(* Logix 5000 project; controller FV vendor 1 type 14 code 217 rev 31.11; software revision 31.00; part 13 of 63 *)
(* tags used below, declared in another part *)
   CWD : CHECKWORD_FLAGS;
   FR_B240 : INT[255];   // DEBOUNCE Debounce Flags
   FR_B246 : INT[255];   // V_REVERSE Flags for reversing contol action
   FR_B3 : INT[255];   // BINARY
   FR_FV29_AV01 : PlantItem;   // FV29_AV01
   FR_FV29_AV04 : PlantItem;   // FV29_AV04
   FR_FV29_AV05 : PlantItem;   // FV29_AV05
   FR_FV29_AV06 : PlantItem;   // FV29_AV06
   FR_FV29_AV07 : PlantItem;   // FV29_AV07
   FR_FV29_ROTO : PlantItem;   // FV29_ROTO
   FR_FV29_VA01 : PlantItem;   // FV29_VA01
   FR_FV30_AV01 : PlantItem;   // FV30_AV01
   FR_FV30_AV04 : PlantItem;   // FV30_AV04
   FR_FV30_AV05 : PlantItem;   // FV30_AV05
   FR_FV30_AV06 : PlantItem;   // FV30_AV06
   FR_FV30_AV07 : PlantItem;   // FV30_AV07
   FR_FV30_ROTO : PlantItem;   // FV30_ROTO
   FR_FV30_VA01 : PlantItem;   // FV30_VA01
   FR_N10 : INT[265];   // FV_AGING Comms to FV Aging PL C
   FR_N100 : INT[265];   // FV FILLING
   FR_N110 : INT[265];   // GREEN BEER Green Beer Main
   FR_N120 : INT[265];   // YEAST CROP Yeast Cropping Main
   FR_N13 : INT[265];   // MV_ROUTE Comms to MV Routing PLC
   FR_N130 : INT[265];   // FILTRATE Filtrate Return
   FR_N14 : INT[265];   // MVFV CIP Comms to MVFV CIP Un it PLC
   FR_N160 : INT[265];   // VESSEL Vessel Working Direc tory
   FR_N200 : INT[265];   // ANALOG_IN Analog Inputs
   FR_N255 : INT[265];   // CHECKWORDS
   FR_N29 : INT[265];   // FV29
   FR_N30 : INT[265];   // FV30
   FR_N7 : INT[265];   // INTEGER
   FR_N99 : INT[265];   // COMMENT Comment Lines
   FR_T144 : TIMER[255];   // CIP
   FR_T4 : TIMER[255];   // TIMER
   FR_T50 : TIMER[52];
   FR_T51 : TIMER[52];
   FR_T52 : TIMER[52];
   FR_T53 : TIMER[52];
   FR_VB1_AV08 : PlantItem;   // VB1_AV08
   FR_VB1_AV09 : PlantItem;   // VB1_AV09
   FR_VB2_AV04 : PlantItem;   // VB2_AV04
   FR_VB2_AV05 : PlantItem;   // VB2_AV05
   FR_VB3_AV04 : PlantItem;   // VB3_AV04
   FR_VB3_AV05 : PlantItem;   // VB3_AV05
   FR_VB4_AV04 : PlantItem;   // VB4_AV04
   FR_VB4_AV05 : PlantItem;   // VB4_AV05
   FR_VB4_AV10 : PlantItem;   // VB4_AV10
   FR_VB4_AV11 : PlantItem;   // VB4_AV11
   FR_VB4_AV16 : PlantItem;   // VB4_AV16
   FR_VB4_AV17 : PlantItem;   // VB4_AV17
(* FR_Common, continued *)

ROUTINE FR_FV29_29   (* ladder *)
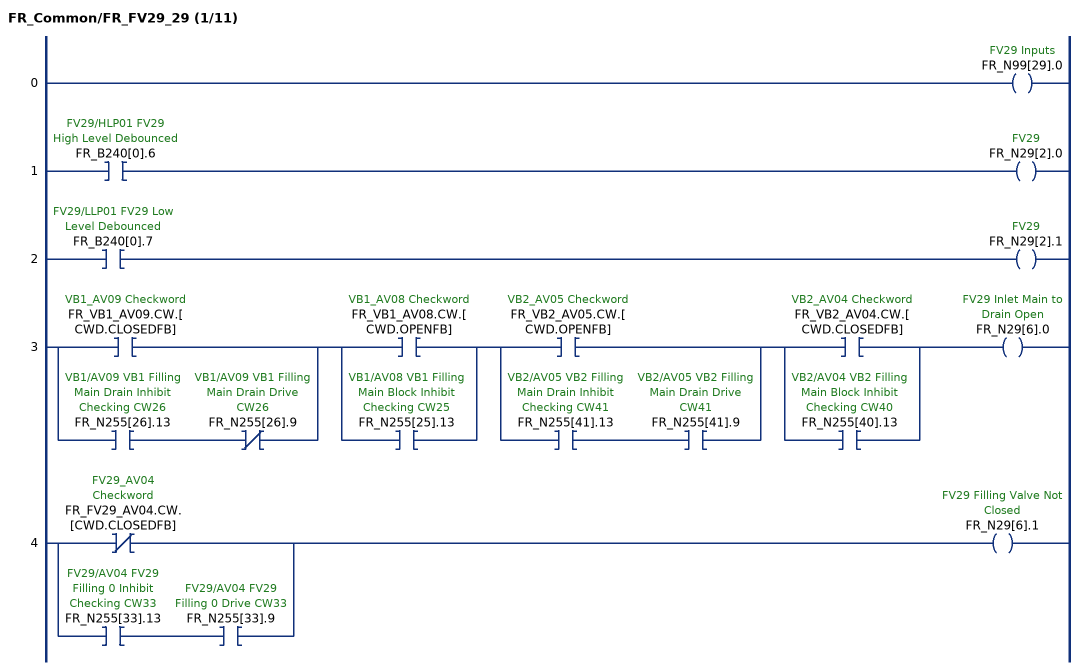
   0: OTE(FR_N99[29].0);
   1: XIC(FR_B240[0].6)OTE(FR_N29[2].0);
   2: XIC(FR_B240[0].7)OTE(FR_N29[2].1);
   3: [XIC(FR_VB1_AV09.CW.[CWD.CLOSEDFB]) ,XIC(FR_N255[26].13) XIO(FR_N255[26].9) ][XIC(FR_VB1_AV08.CW.[CWD.OPENFB]) ,XIC(FR_N255[25].13) ][XIC(FR_VB2_AV05.CW.[CWD.OPENFB]) ,XIC(FR_N255[41].13) XIC(FR_N255[41].9) ][XIC(FR_VB2_AV04.CW.[CWD.CLOSEDFB]) ,XIC(FR_N255[40].13) ]OTE(FR_N29[6].0);
   4: [XIO(FR_FV29_AV04.CW.[CWD.CLOSEDFB]) ,XIC(FR_N255[33].13) XIC(FR_N255[33].9) ]OTE(FR_N29[6].1);
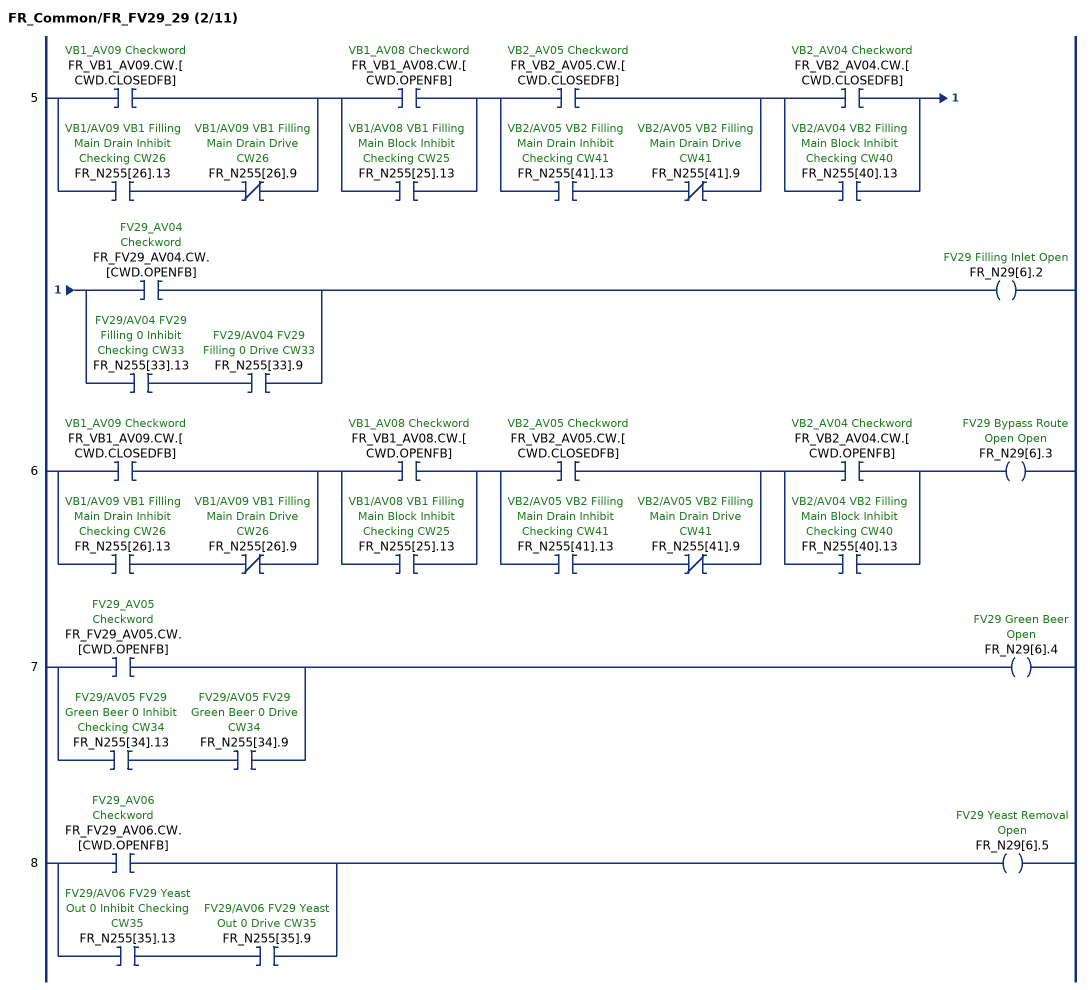
   5: [XIC(FR_VB1_AV09.CW.[CWD.CLOSEDFB]) ,XIC(FR_N255[26].13) XIO(FR_N255[26].9) ][XIC(FR_VB1_AV08.CW.[CWD.OPENFB]) ,XIC(FR_N255[25].13) ][XIC(FR_VB2_AV05.CW.[CWD.CLOSEDFB]) ,XIC(FR_N255[41].13) XIO(FR_N255[41].9) ][XIC(FR_VB2_AV04.CW.[CWD.CLOSEDFB]) ,XIC(FR_N255[40].13) ][XIC(FR_FV29_AV04.CW.[CWD.OPENFB]) ,XIC(FR_N255[33].13) XIC(FR_N255[33].9) ]OTE(FR_N29[6].2);
   6: [XIC(FR_VB1_AV09.CW.[CWD.CLOSEDFB]) ,XIC(FR_N255[26].13) XIO(FR_N255[26].9) ][XIC(FR_VB1_AV08.CW.[CWD.OPENFB]) ,XIC(FR_N255[25].13) ][XIC(FR_VB2_AV05.CW.[CWD.CLOSEDFB]) ,XIC(FR_N255[41].13) XIO(FR_N255[41].9) ][XIC(FR_VB2_AV04.CW.[CWD.OPENFB]) ,XIC(FR_N255[40].13) ]OTE(FR_N29[6].3);
   7: [XIC(FR_FV29_AV05.CW.[CWD.OPENFB]) ,XIC(FR_N255[34].13) XIC(FR_N255[34].9) ]OTE(FR_N29[6].4);
   8: [XIC(FR_FV29_AV06.CW.[CWD.OPENFB]) ,XIC(FR_N255[35].13) XIC(FR_N255[35].9) ]OTE(FR_N29[6].5);
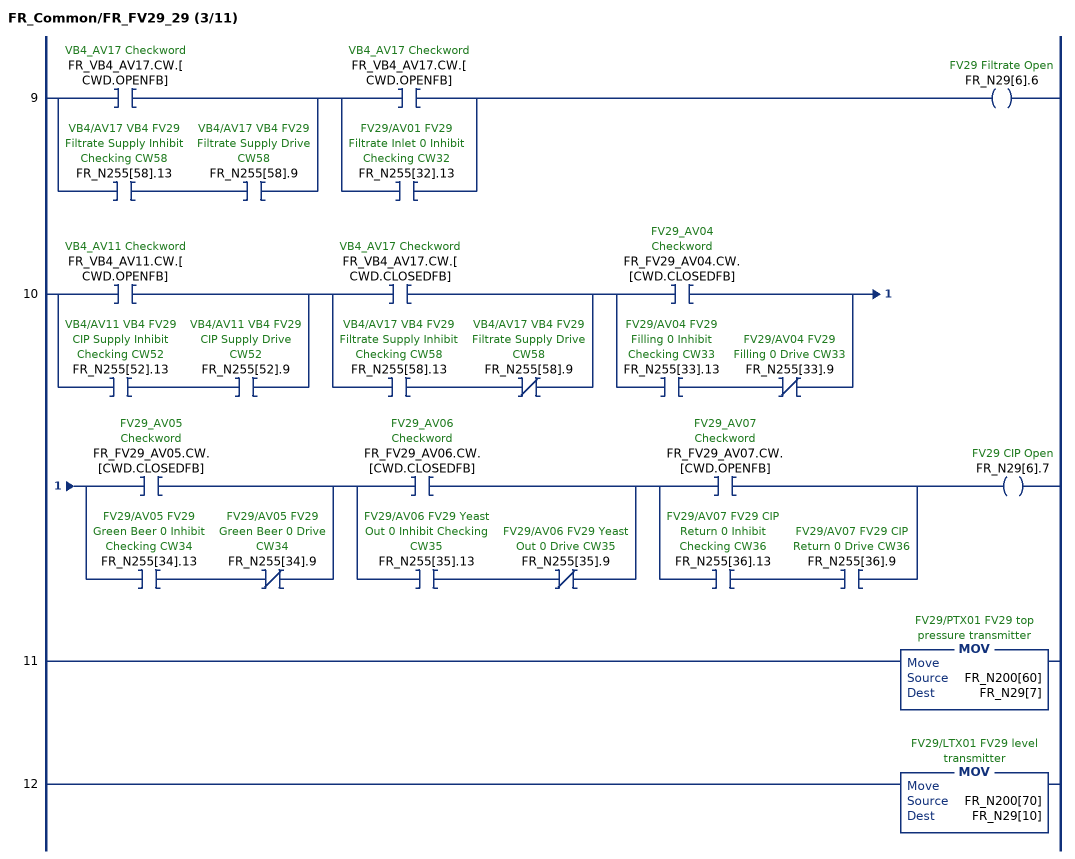
   9: [XIC(FR_VB4_AV17.CW.[CWD.OPENFB]) ,XIC(FR_N255[58].13) XIC(FR_N255[58].9) ][XIC(FR_VB4_AV17.CW.[CWD.OPENFB]) ,XIC(FR_N255[32].13) ]OTE(FR_N29[6].6);
   10: [XIC(FR_VB4_AV11.CW.[CWD.OPENFB]) ,XIC(FR_N255[52].13) XIC(FR_N255[52].9) ][XIC(FR_VB4_AV17.CW.[CWD.CLOSEDFB]) ,XIC(FR_N255[58].13) XIO(FR_N255[58].9) ][XIC(FR_FV29_AV04.CW.[CWD.CLOSEDFB]) ,XIC(FR_N255[33].13) XIO(FR_N255[33].9) ][XIC(FR_FV29_AV05.CW.[CWD.CLOSEDFB]) ,XIC(FR_N255[34].13) XIO(FR_N255[34].9) ][XIC(FR_FV29_AV06.CW.[CWD.CLOSEDFB]) ,XIC(FR_N255[35].13) XIO(FR_N255[35].9) ][XIC(FR_FV29_AV07.CW.[CWD.OPENFB]) ,XIC(FR_N255[36].13) XIC(FR_N255[36].9) ]OTE(FR_N29[6].7);
   11: MOV(FR_N200[60],FR_N29[7]);
   12: MOV(FR_N200[70],FR_N29[10]);
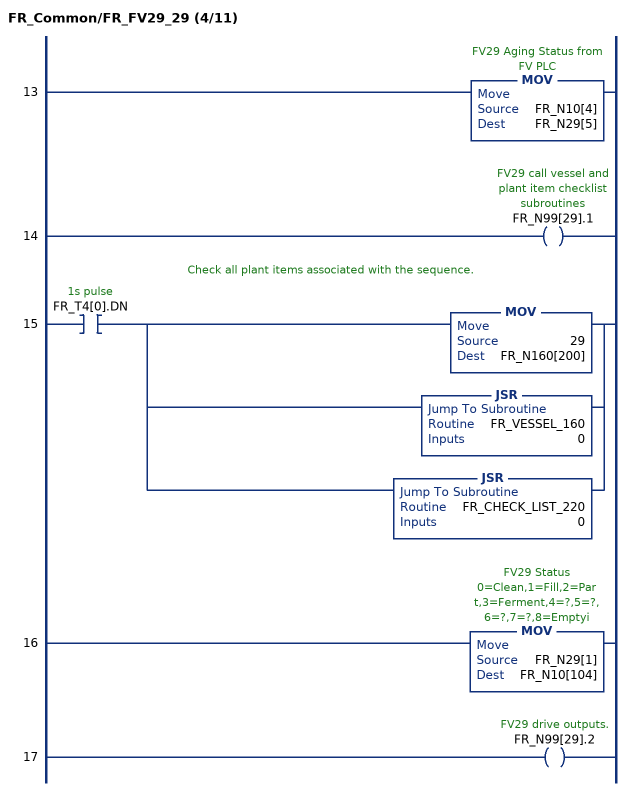
   13: MOV(FR_N10[4],FR_N29[5]);
   14: OTE(FR_N99[29].1);
   // Check all plant items associated with the sequence.
   15: XIC(FR_T4[0].DN)[MOV(29,FR_N160[200]) ,JSR(FR_VESSEL_160,0) ,JSR(FR_CHECK_LIST_220,0) ];
   16: MOV(FR_N29[1],FR_N10[104]);
   17: OTE(FR_N99[29].2);
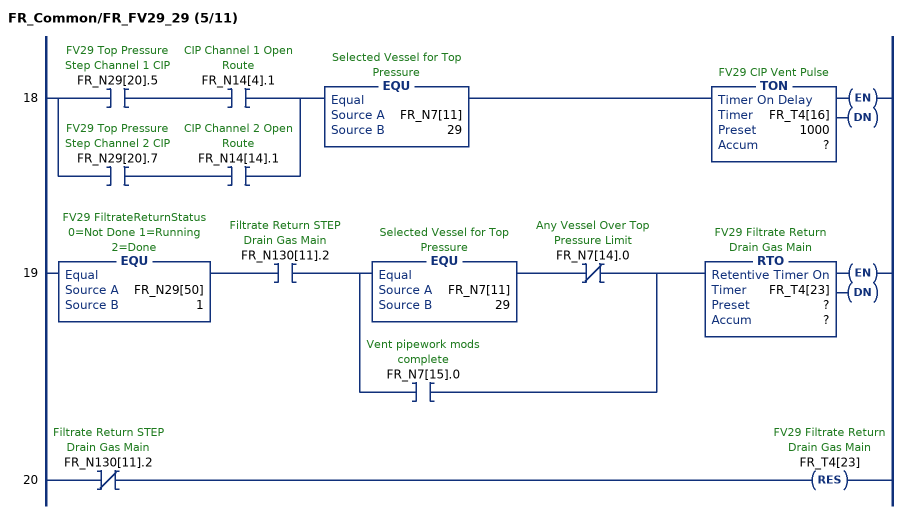
   18: [XIC(FR_N29[20].5) XIC(FR_N14[4].1) ,XIC(FR_N29[20].7) XIC(FR_N14[14].1) ]EQU(FR_N7[11],29)TON(FR_T4[16],?,?);
   19: EQU(FR_N29[50],1)XIC(FR_N130[11].2)[EQU(FR_N7[11],29) XIO(FR_N7[14].0) ,XIC(FR_N7[15].0) ]RTO(FR_T4[23],?,?);
   20: XIO(FR_N130[11].2)RES(FR_T4[23]);
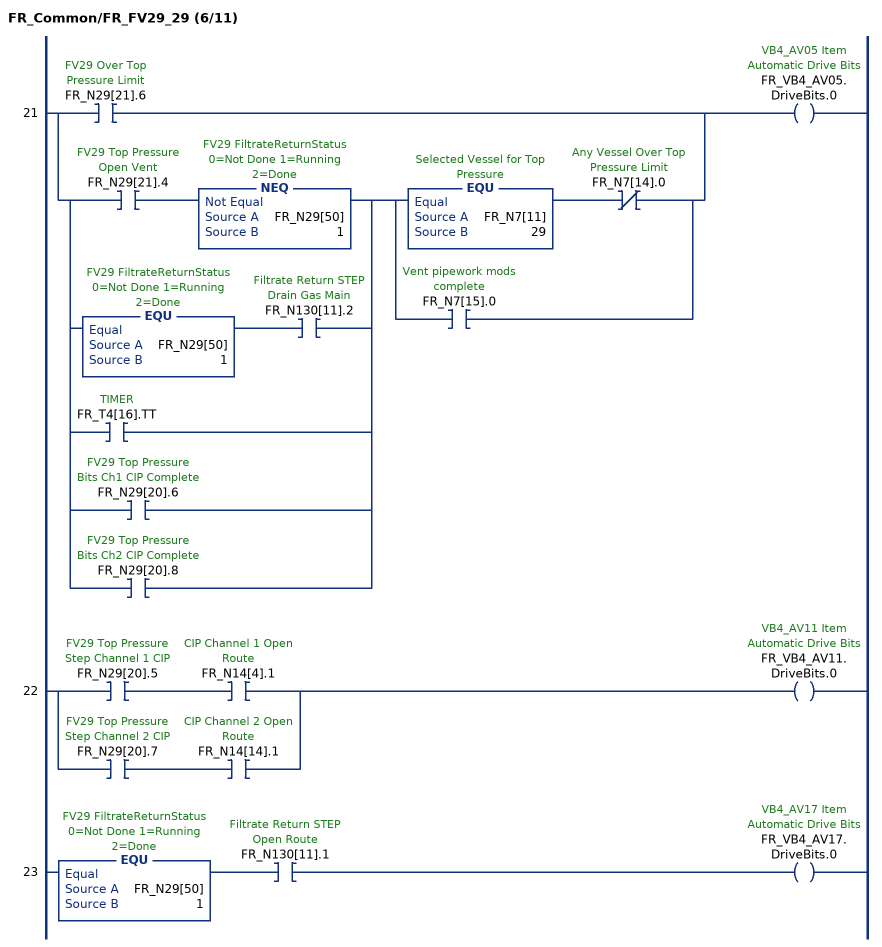
   21: [XIC(FR_N29[21].6) ,[XIC(FR_N29[21].4) NEQ(FR_N29[50],1) ,EQU(FR_N29[50],1) XIC(FR_N130[11].2) ,XIC(FR_T4[16].TT) ,[XIC(FR_N29[20].6) ,XIC(FR_N29[20].8) ] ] [EQU(FR_N7[11],29) XIO(FR_N7[14].0) ,XIC(FR_N7[15].0) ] ]OTE(FR_VB4_AV05.DriveBits.0);
   22: [XIC(FR_N29[20].5) XIC(FR_N14[4].1) ,XIC(FR_N29[20].7) XIC(FR_N14[14].1) ]OTE(FR_VB4_AV11.DriveBits.0);
   23: EQU(FR_N29[50],1)XIC(FR_N130[11].1)OTE(FR_VB4_AV17.DriveBits.0);
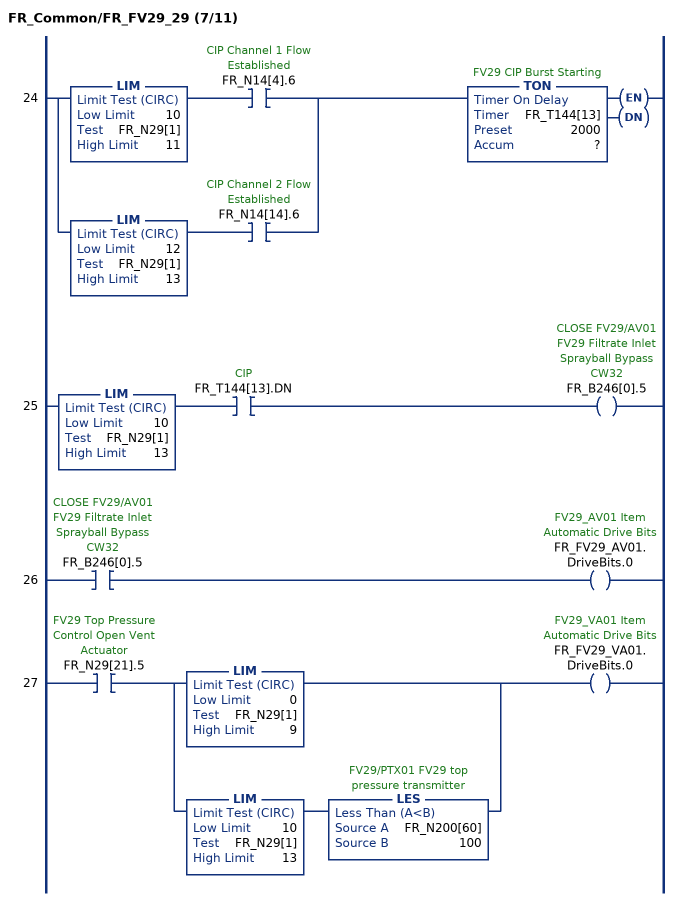
   24: [LIM(10,FR_N29[1],11) XIC(FR_N14[4].6) ,LIM(12,FR_N29[1],13) XIC(FR_N14[14].6) ]TON(FR_T144[13],?,?);
   25: LIM(10,FR_N29[1],13)XIC(FR_T144[13].DN)OTE(FR_B246[0].5);
   26: XIC(FR_B246[0].5)OTE(FR_FV29_AV01.DriveBits.0);
   27: XIC(FR_N29[21].5)[LIM(0,FR_N29[1],9) ,LIM(10,FR_N29[1],13) LES(FR_N200[60],100) ]OTE(FR_FV29_VA01.DriveBits.0);
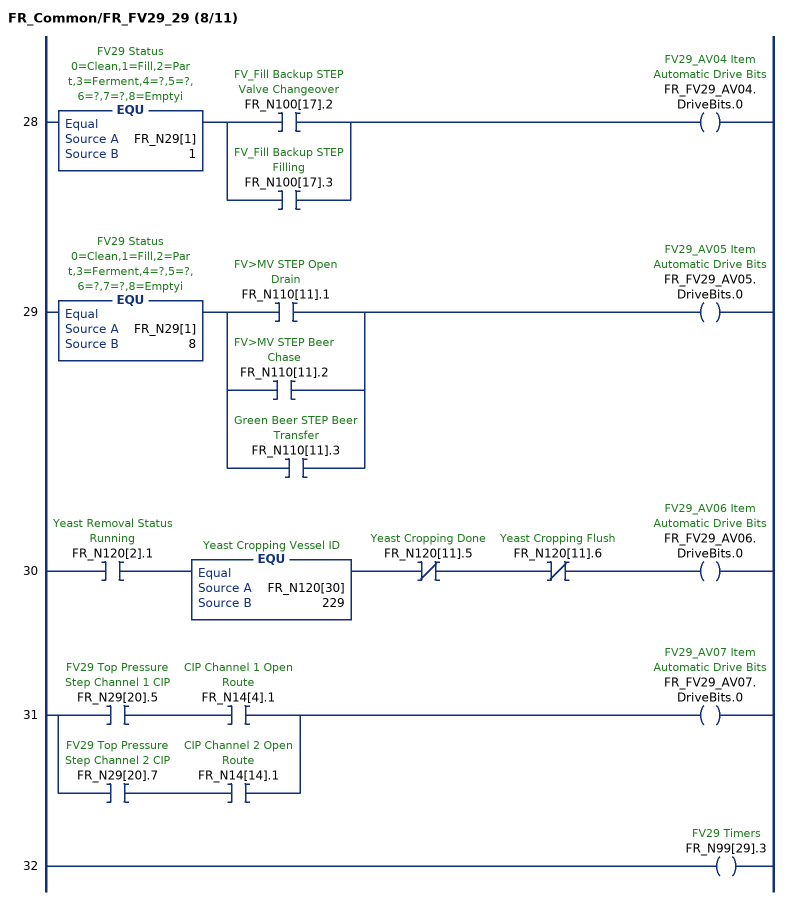
   28: EQU(FR_N29[1],1)[XIC(FR_N100[17].2) ,XIC(FR_N100[17].3) ]OTE(FR_FV29_AV04.DriveBits.0);
   29: EQU(FR_N29[1],8)[XIC(FR_N110[11].1) ,XIC(FR_N110[11].2) ,XIC(FR_N110[11].3) ]OTE(FR_FV29_AV05.DriveBits.0);
   30: XIC(FR_N120[2].1)EQU(FR_N120[30],229)XIO(FR_N120[11].5)XIO(FR_N120[11].6)OTE(FR_FV29_AV06.DriveBits.0);
   31: [XIC(FR_N29[20].5) XIC(FR_N14[4].1) ,XIC(FR_N29[20].7) XIC(FR_N14[14].1) ]OTE(FR_FV29_AV07.DriveBits.0);
   32: OTE(FR_N99[29].3);
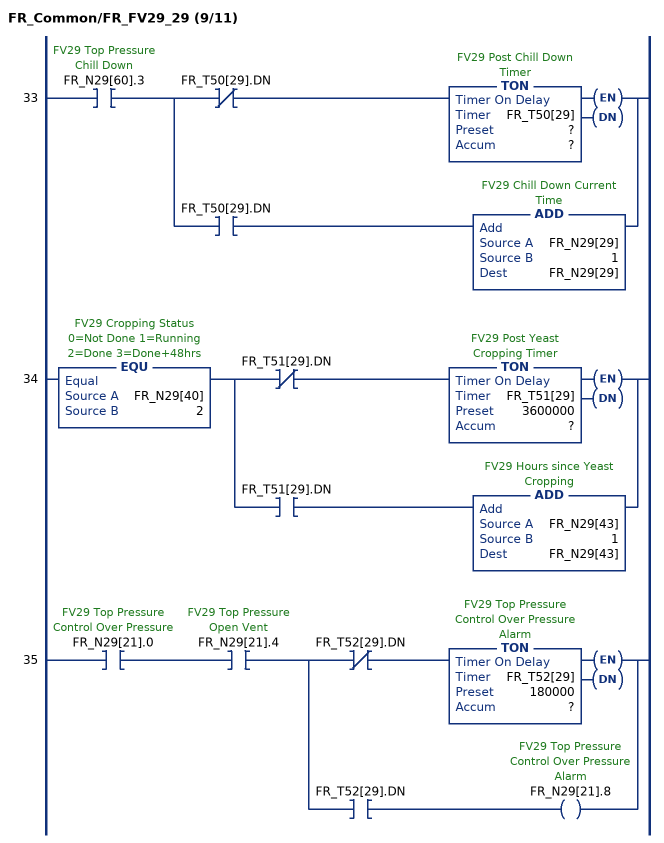
   33: XIC(FR_N29[60].3)[XIO(FR_T50[29].DN) TON(FR_T50[29],?,?) ,XIC(FR_T50[29].DN) ADD(FR_N29[29],1,FR_N29[29]) ];
   34: EQU(FR_N29[40],2)[XIO(FR_T51[29].DN) TON(FR_T51[29],?,?) ,XIC(FR_T51[29].DN) ADD(FR_N29[43],1,FR_N29[43]) ];
   35: XIC(FR_N29[21].0)XIC(FR_N29[21].4)[XIO(FR_T52[29].DN) TON(FR_T52[29],?,?) ,XIC(FR_T52[29].DN) OTE(FR_N29[21].8) ];
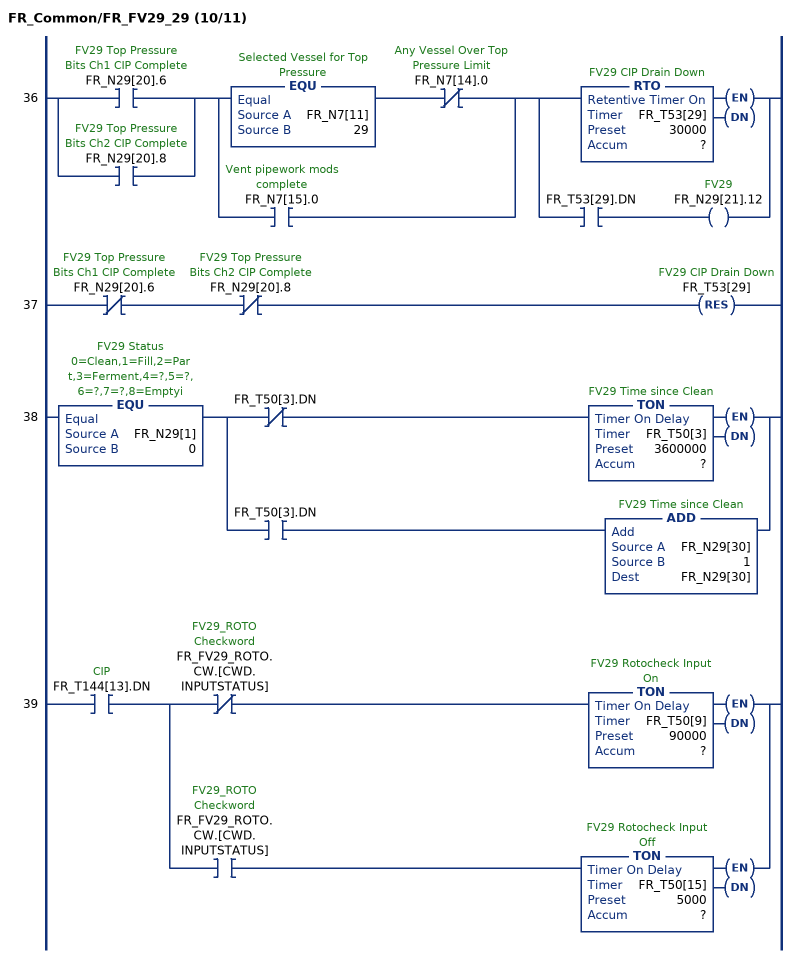
   36: [XIC(FR_N29[20].6) ,XIC(FR_N29[20].8) ][EQU(FR_N7[11],29) XIO(FR_N7[14].0) ,XIC(FR_N7[15].0) ][RTO(FR_T53[29],?,?) ,XIC(FR_T53[29].DN) OTE(FR_N29[21].12) ];
   37: XIO(FR_N29[20].6)XIO(FR_N29[20].8)RES(FR_T53[29]);
   38: EQU(FR_N29[1],0)[XIO(FR_T50[3].DN) TON(FR_T50[3],?,?) ,XIC(FR_T50[3].DN) ADD(FR_N29[30],1,FR_N29[30]) ];
   39: XIC(FR_T144[13].DN)[XIO(FR_FV29_ROTO.CW.[CWD.INPUTSTATUS]) TON(FR_T50[9],?,?) ,XIC(FR_FV29_ROTO.CW.[CWD.INPUTSTATUS]) TON(FR_T50[15],?,?) ];
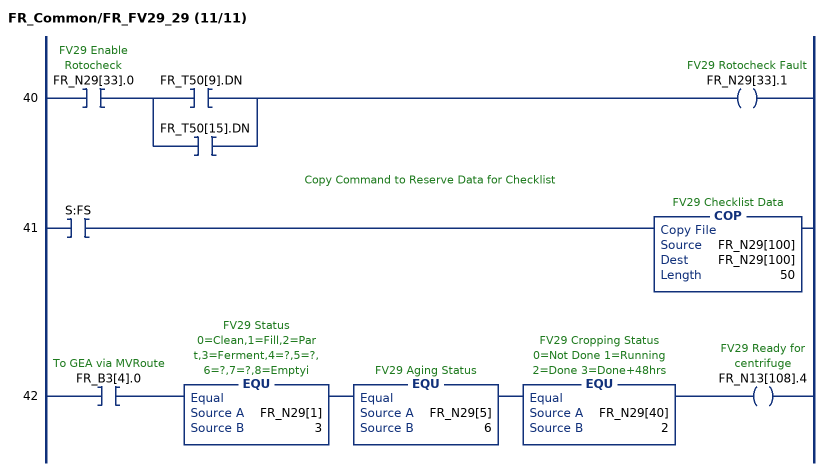
   40: XIC(FR_N29[33].0)[XIC(FR_T50[9].DN) ,XIC(FR_T50[15].DN) ]OTE(FR_N29[33].1);
   // Copy Command to Reserve Data for Checklist
   41: XIC(S:FS)COP(FR_N29[100],FR_N29[100],50);
   42: XIC(FR_B3[4].0)EQU(FR_N29[1],3)EQU(FR_N29[5],6)EQU(FR_N29[40],2)OTE(FR_N13[108].4);
END_ROUTINE

ROUTINE FR_FV30_30   (* ladder *)
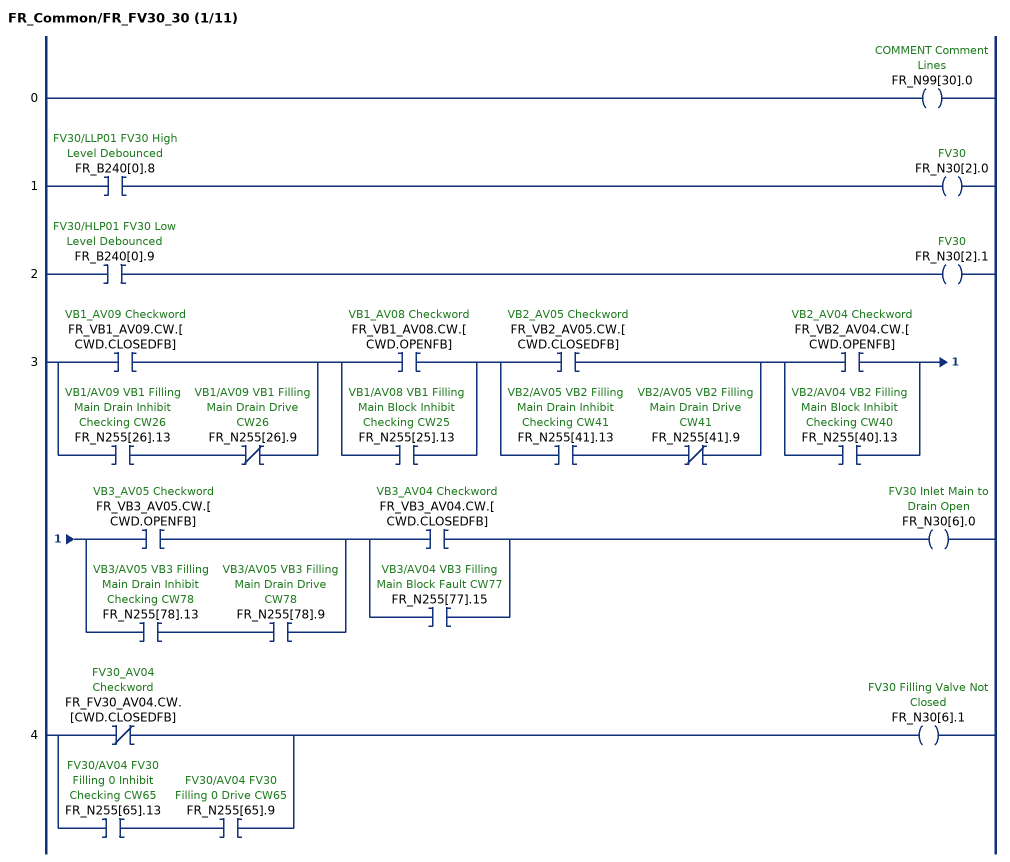
   0: OTE(FR_N99[30].0);
   1: XIC(FR_B240[0].8)OTE(FR_N30[2].0);
   2: XIC(FR_B240[0].9)OTE(FR_N30[2].1);
   3: [XIC(FR_VB1_AV09.CW.[CWD.CLOSEDFB]) ,XIC(FR_N255[26].13) XIO(FR_N255[26].9) ][XIC(FR_VB1_AV08.CW.[CWD.OPENFB]) ,XIC(FR_N255[25].13) ][XIC(FR_VB2_AV05.CW.[CWD.CLOSEDFB]) ,XIC(FR_N255[41].13) XIO(FR_N255[41].9) ][XIC(FR_VB2_AV04.CW.[CWD.OPENFB]) ,XIC(FR_N255[40].13) ][XIC(FR_VB3_AV05.CW.[CWD.OPENFB]) ,XIC(FR_N255[78].13) XIC(FR_N255[78].9) ][XIC(FR_VB3_AV04.CW.[CWD.CLOSEDFB]) ,XIC(FR_N255[77].15) ]OTE(FR_N30[6].0);
   4: [XIO(FR_FV30_AV04.CW.[CWD.CLOSEDFB]) ,XIC(FR_N255[65].13) XIC(FR_N255[65].9) ]OTE(FR_N30[6].1);
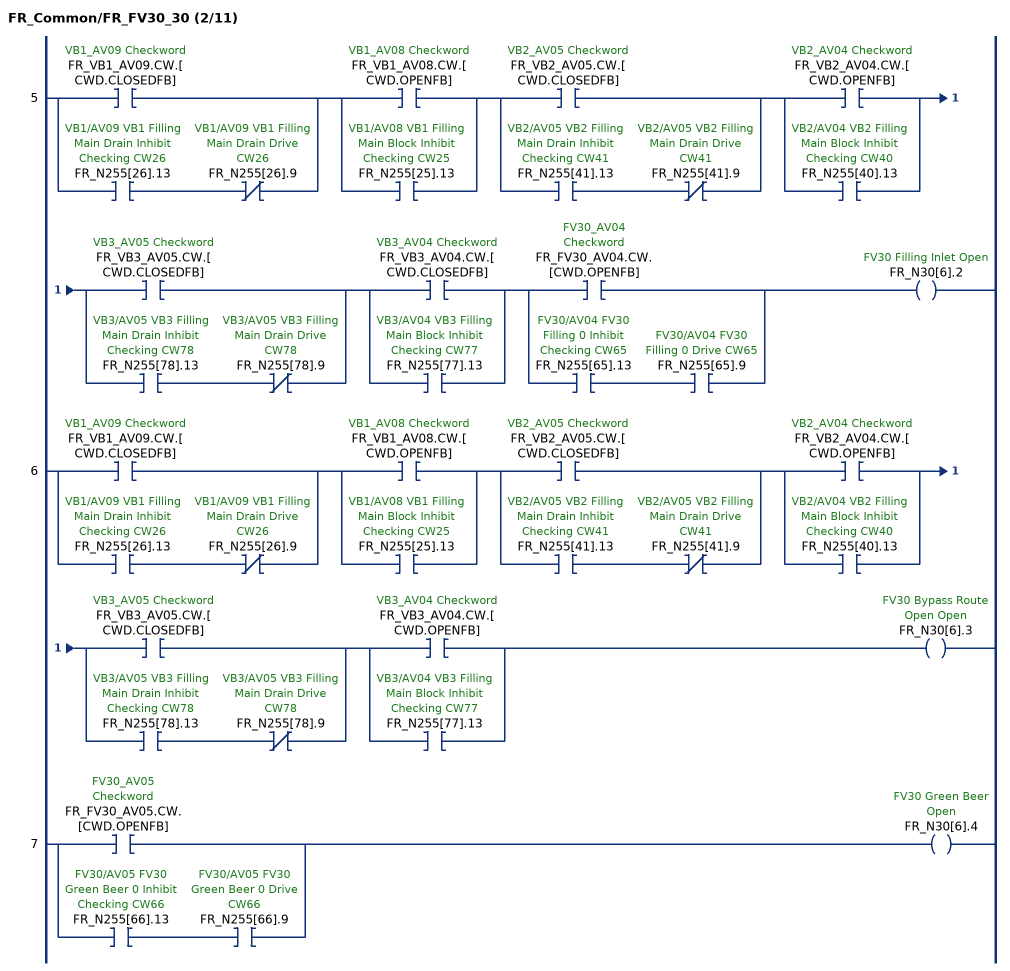
   5: [XIC(FR_VB1_AV09.CW.[CWD.CLOSEDFB]) ,XIC(FR_N255[26].13) XIO(FR_N255[26].9) ][XIC(FR_VB1_AV08.CW.[CWD.OPENFB]) ,XIC(FR_N255[25].13) ][XIC(FR_VB2_AV05.CW.[CWD.CLOSEDFB]) ,XIC(FR_N255[41].13) XIO(FR_N255[41].9) ][XIC(FR_VB2_AV04.CW.[CWD.OPENFB]) ,XIC(FR_N255[40].13) ][XIC(FR_VB3_AV05.CW.[CWD.CLOSEDFB]) ,XIC(FR_N255[78].13) XIO(FR_N255[78].9) ][XIC(FR_VB3_AV04.CW.[CWD.CLOSEDFB]) ,XIC(FR_N255[77].13) ][XIC(FR_FV30_AV04.CW.[CWD.OPENFB]) ,XIC(FR_N255[65].13) XIC(FR_N255[65].9) ]OTE(FR_N30[6].2);
   6: [XIC(FR_VB1_AV09.CW.[CWD.CLOSEDFB]) ,XIC(FR_N255[26].13) XIO(FR_N255[26].9) ][XIC(FR_VB1_AV08.CW.[CWD.OPENFB]) ,XIC(FR_N255[25].13) ][XIC(FR_VB2_AV05.CW.[CWD.CLOSEDFB]) ,XIC(FR_N255[41].13) XIO(FR_N255[41].9) ][XIC(FR_VB2_AV04.CW.[CWD.OPENFB]) ,XIC(FR_N255[40].13) ][XIC(FR_VB3_AV05.CW.[CWD.CLOSEDFB]) ,XIC(FR_N255[78].13) XIO(FR_N255[78].9) ][XIC(FR_VB3_AV04.CW.[CWD.OPENFB]) ,XIC(FR_N255[77].13) ]OTE(FR_N30[6].3);
   7: [XIC(FR_FV30_AV05.CW.[CWD.OPENFB]) ,XIC(FR_N255[66].13) XIC(FR_N255[66].9) ]OTE(FR_N30[6].4);
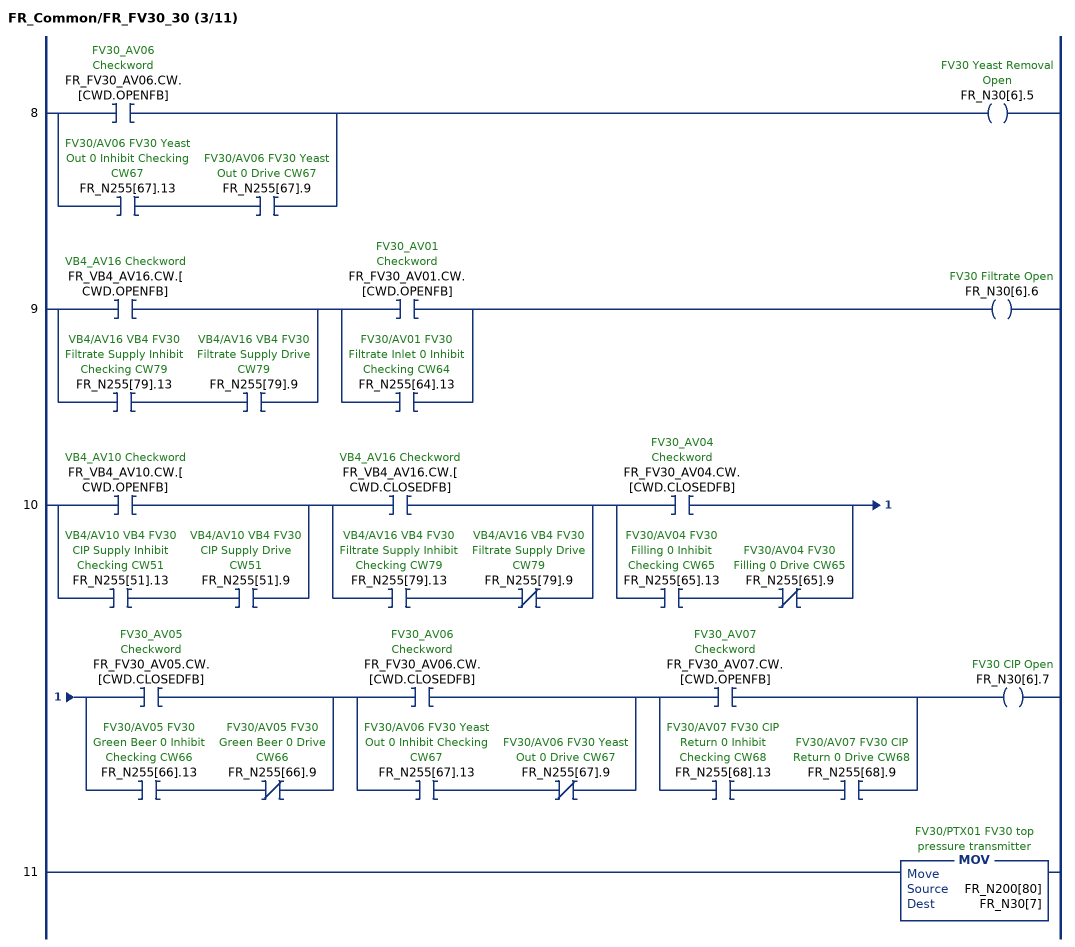
   8: [XIC(FR_FV30_AV06.CW.[CWD.OPENFB]) ,XIC(FR_N255[67].13) XIC(FR_N255[67].9) ]OTE(FR_N30[6].5);
   9: [XIC(FR_VB4_AV16.CW.[CWD.OPENFB]) ,XIC(FR_N255[79].13) XIC(FR_N255[79].9) ][XIC(FR_FV30_AV01.CW.[CWD.OPENFB]) ,XIC(FR_N255[64].13) ]OTE(FR_N30[6].6);
   10: [XIC(FR_VB4_AV10.CW.[CWD.OPENFB]) ,XIC(FR_N255[51].13) XIC(FR_N255[51].9) ][XIC(FR_VB4_AV16.CW.[CWD.CLOSEDFB]) ,XIC(FR_N255[79].13) XIO(FR_N255[79].9) ][XIC(FR_FV30_AV04.CW.[CWD.CLOSEDFB]) ,XIC(FR_N255[65].13) XIO(FR_N255[65].9) ][XIC(FR_FV30_AV05.CW.[CWD.CLOSEDFB]) ,XIC(FR_N255[66].13) XIO(FR_N255[66].9) ][XIC(FR_FV30_AV06.CW.[CWD.CLOSEDFB]) ,XIC(FR_N255[67].13) XIO(FR_N255[67].9) ][XIC(FR_FV30_AV07.CW.[CWD.OPENFB]) ,XIC(FR_N255[68].13) XIC(FR_N255[68].9) ]OTE(FR_N30[6].7);
   11: MOV(FR_N200[80],FR_N30[7]);
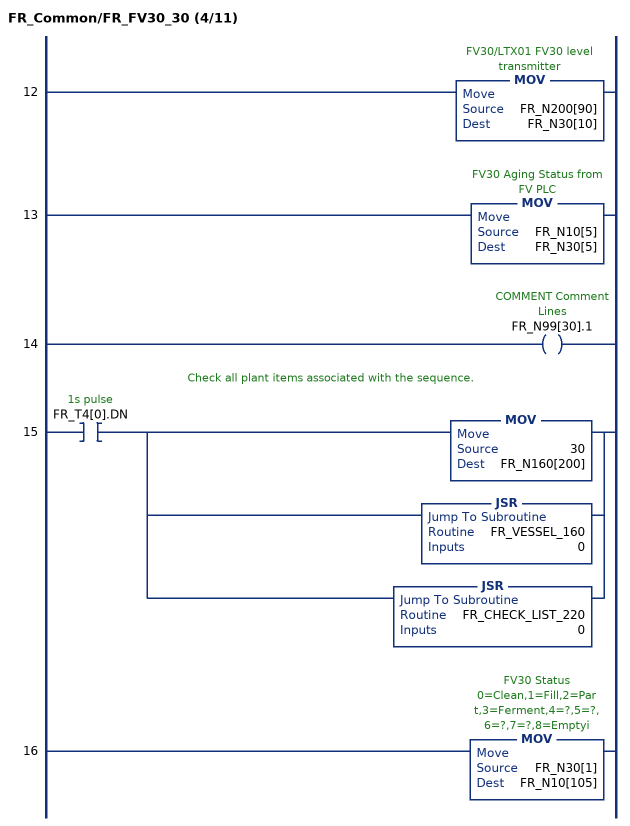
   12: MOV(FR_N200[90],FR_N30[10]);
   13: MOV(FR_N10[5],FR_N30[5]);
   14: OTE(FR_N99[30].1);
   // Check all plant items associated with the sequence.
   15: XIC(FR_T4[0].DN)[MOV(30,FR_N160[200]) ,JSR(FR_VESSEL_160,0) ,JSR(FR_CHECK_LIST_220,0) ];
   16: MOV(FR_N30[1],FR_N10[105]);
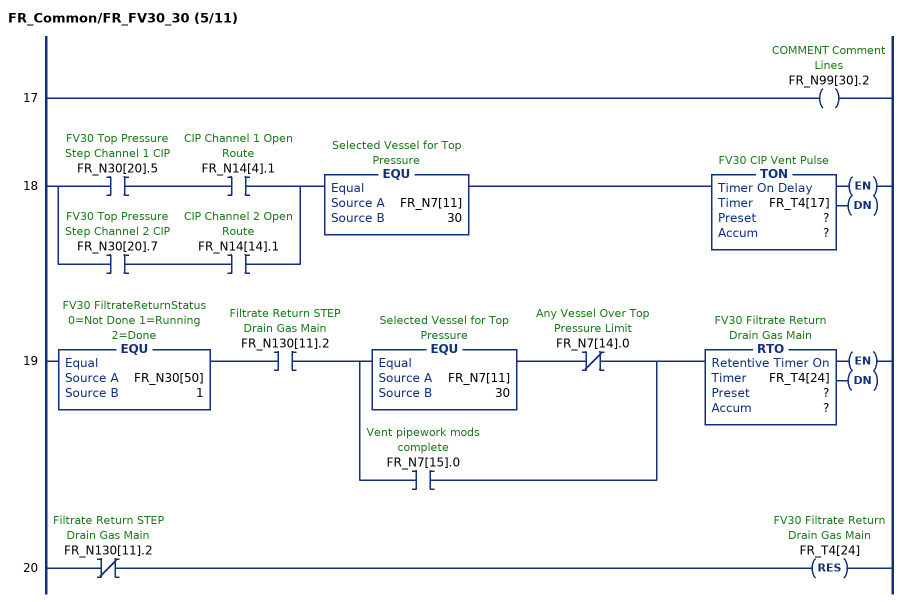
   17: OTE(FR_N99[30].2);
   18: [XIC(FR_N30[20].5) XIC(FR_N14[4].1) ,XIC(FR_N30[20].7) XIC(FR_N14[14].1) ]EQU(FR_N7[11],30)TON(FR_T4[17],?,?);
   19: EQU(FR_N30[50],1)XIC(FR_N130[11].2)[EQU(FR_N7[11],30) XIO(FR_N7[14].0) ,XIC(FR_N7[15].0) ]RTO(FR_T4[24],?,?);
   20: XIO(FR_N130[11].2)RES(FR_T4[24]);
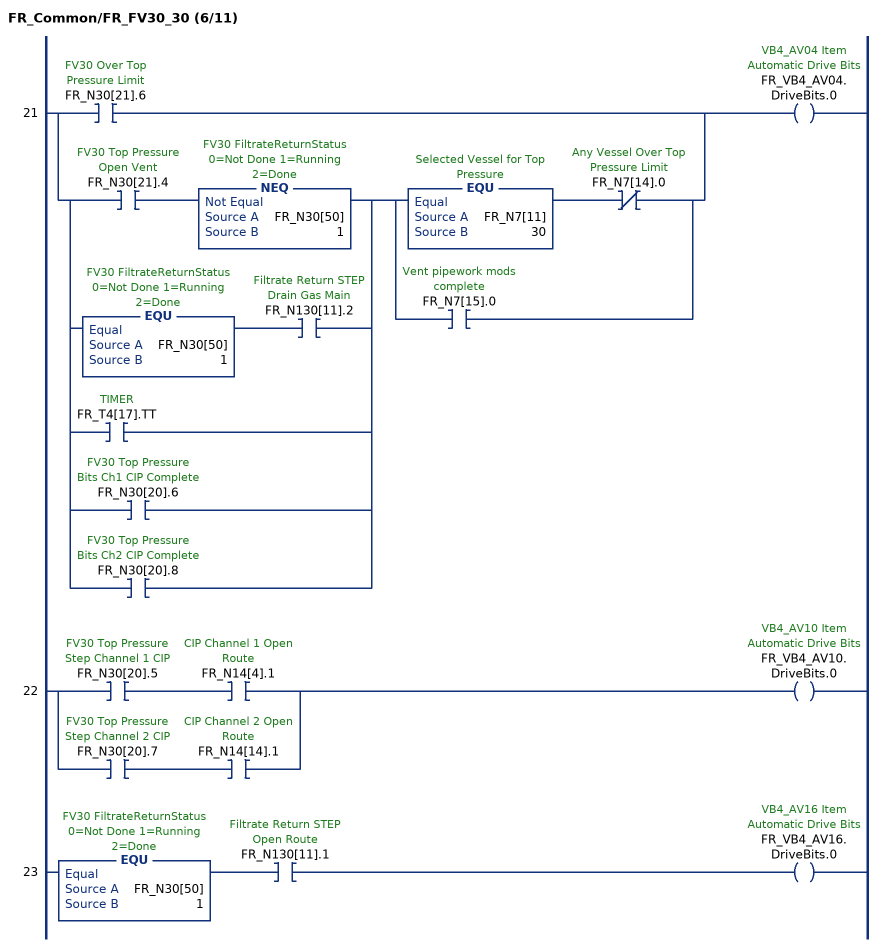
   21: [XIC(FR_N30[21].6) ,[XIC(FR_N30[21].4) NEQ(FR_N30[50],1) ,EQU(FR_N30[50],1) XIC(FR_N130[11].2) ,XIC(FR_T4[17].TT) ,[XIC(FR_N30[20].6) ,XIC(FR_N30[20].8) ] ] [EQU(FR_N7[11],30) XIO(FR_N7[14].0) ,XIC(FR_N7[15].0) ] ]OTE(FR_VB4_AV04.DriveBits.0);
   22: [XIC(FR_N30[20].5) XIC(FR_N14[4].1) ,XIC(FR_N30[20].7) XIC(FR_N14[14].1) ]OTE(FR_VB4_AV10.DriveBits.0);
   23: EQU(FR_N30[50],1)XIC(FR_N130[11].1)OTE(FR_VB4_AV16.DriveBits.0);
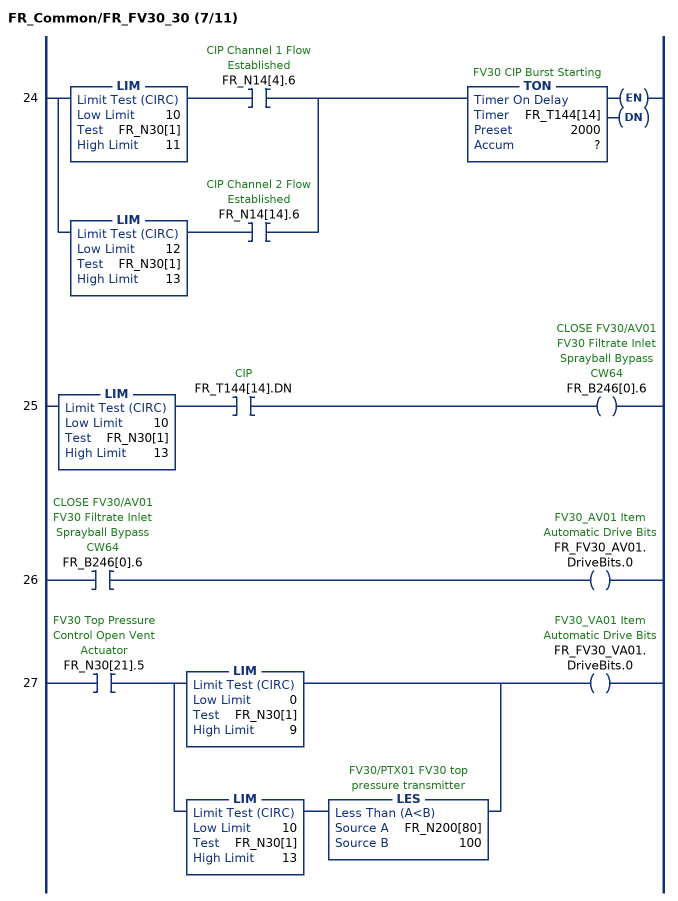
   24: [LIM(10,FR_N30[1],11) XIC(FR_N14[4].6) ,LIM(12,FR_N30[1],13) XIC(FR_N14[14].6) ]TON(FR_T144[14],?,?);
   25: LIM(10,FR_N30[1],13)XIC(FR_T144[14].DN)OTE(FR_B246[0].6);
   26: XIC(FR_B246[0].6)OTE(FR_FV30_AV01.DriveBits.0);
   27: XIC(FR_N30[21].5)[LIM(0,FR_N30[1],9) ,LIM(10,FR_N30[1],13) LES(FR_N200[80],100) ]OTE(FR_FV30_VA01.DriveBits.0);
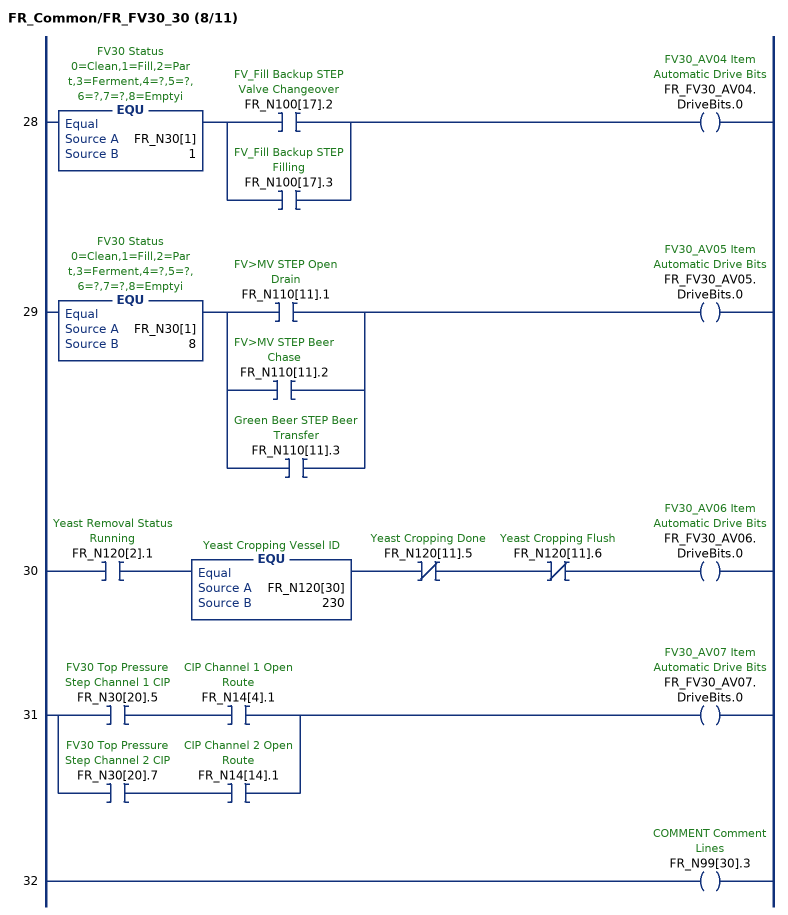
   28: EQU(FR_N30[1],1)[XIC(FR_N100[17].2) ,XIC(FR_N100[17].3) ]OTE(FR_FV30_AV04.DriveBits.0);
   29: EQU(FR_N30[1],8)[XIC(FR_N110[11].1) ,XIC(FR_N110[11].2) ,XIC(FR_N110[11].3) ]OTE(FR_FV30_AV05.DriveBits.0);
   30: XIC(FR_N120[2].1)EQU(FR_N120[30],230)XIO(FR_N120[11].5)XIO(FR_N120[11].6)OTE(FR_FV30_AV06.DriveBits.0);
   31: [XIC(FR_N30[20].5) XIC(FR_N14[4].1) ,XIC(FR_N30[20].7) XIC(FR_N14[14].1) ]OTE(FR_FV30_AV07.DriveBits.0);
   32: OTE(FR_N99[30].3);
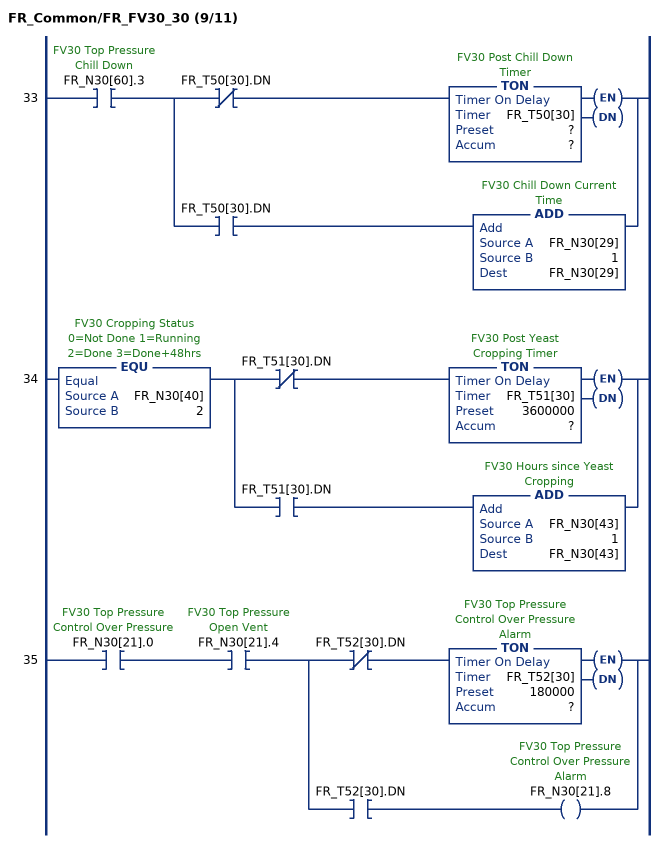
   33: XIC(FR_N30[60].3)[XIO(FR_T50[30].DN) TON(FR_T50[30],?,?) ,XIC(FR_T50[30].DN) ADD(FR_N30[29],1,FR_N30[29]) ];
   34: EQU(FR_N30[40],2)[XIO(FR_T51[30].DN) TON(FR_T51[30],?,?) ,XIC(FR_T51[30].DN) ADD(FR_N30[43],1,FR_N30[43]) ];
   35: XIC(FR_N30[21].0)XIC(FR_N30[21].4)[XIO(FR_T52[30].DN) TON(FR_T52[30],?,?) ,XIC(FR_T52[30].DN) OTE(FR_N30[21].8) ];
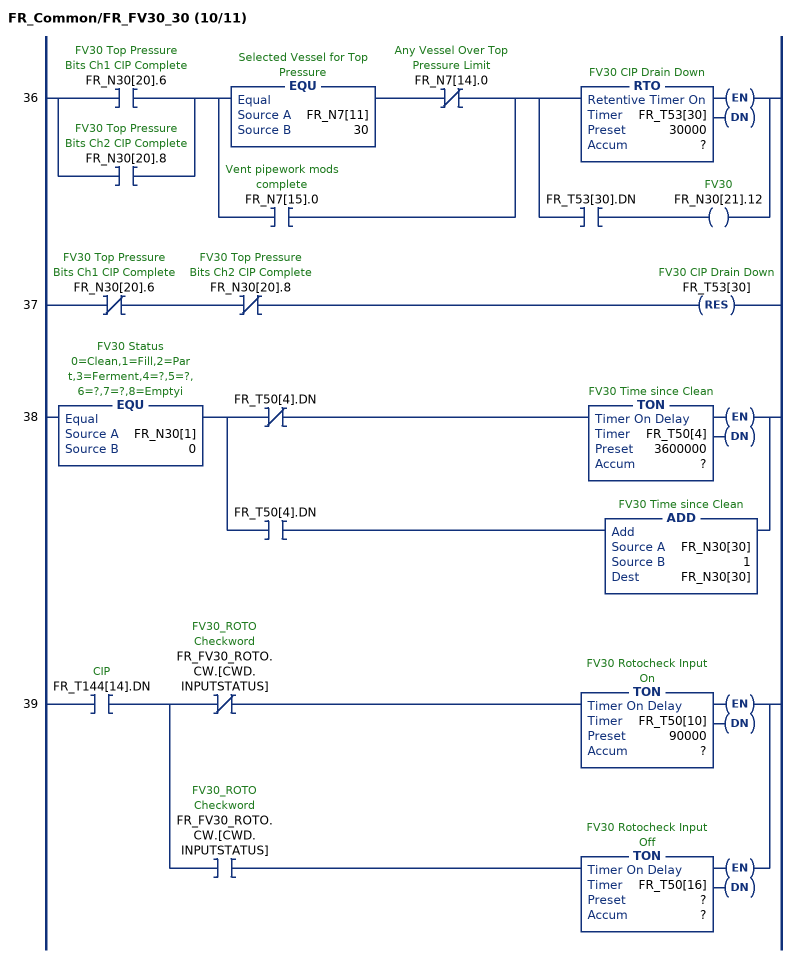
   36: [XIC(FR_N30[20].6) ,XIC(FR_N30[20].8) ][EQU(FR_N7[11],30) XIO(FR_N7[14].0) ,XIC(FR_N7[15].0) ][RTO(FR_T53[30],?,?) ,XIC(FR_T53[30].DN) OTE(FR_N30[21].12) ];
   37: XIO(FR_N30[20].6)XIO(FR_N30[20].8)RES(FR_T53[30]);
   38: EQU(FR_N30[1],0)[XIO(FR_T50[4].DN) TON(FR_T50[4],?,?) ,XIC(FR_T50[4].DN) ADD(FR_N30[30],1,FR_N30[30]) ];
   39: XIC(FR_T144[14].DN)[XIO(FR_FV30_ROTO.CW.[CWD.INPUTSTATUS]) TON(FR_T50[10],?,?) ,XIC(FR_FV30_ROTO.CW.[CWD.INPUTSTATUS]) TON(FR_T50[16],?,?) ];
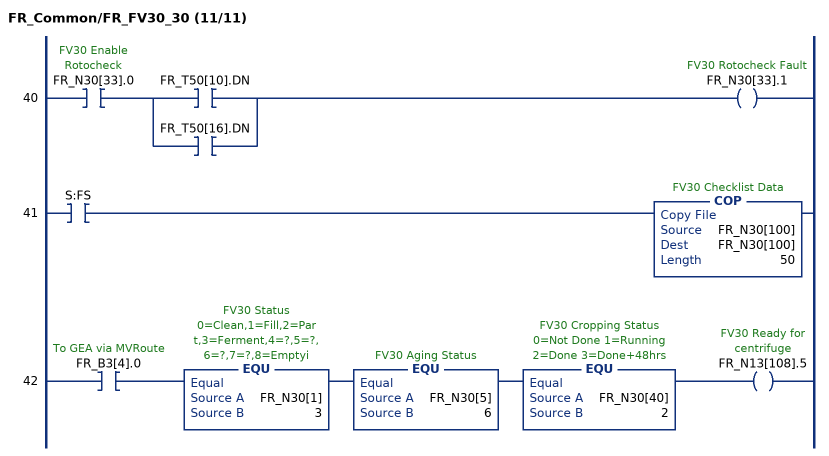
   40: XIC(FR_N30[33].0)[XIC(FR_T50[10].DN) ,XIC(FR_T50[16].DN) ]OTE(FR_N30[33].1);
   41: XIC(S:FS)COP(FR_N30[100],FR_N30[100],50);
   42: XIC(FR_B3[4].0)EQU(FR_N30[1],3)EQU(FR_N30[5],6)EQU(FR_N30[40],2)OTE(FR_N13[108].5);
END_ROUTINE
